screen "BWT Target Setpoints" 1280x800, template "Template"
   on GenerateScreen: "TitleUpdater"()
   Button "HmiScreenItemData_1" at 1,1 size 150x43; TextOn 'Back'; TextOff 'Commissioning'
      on Release: ActivateScreen("Commissioning Main Page", 0)
   AlarmView "Alarm view_1" at 0,777 size 1280x23
   IOField "I/O field_3" at 570,423 size 115x22; FormatPattern 9999.9; Unit Nm³/hr
      ProcessValue <- "2084_Setpoints_FIT420_LoLo"
   TextField "Text field_10" at 47,184 size 216x30; Text 'Description'
   TextField "Text field_6" at 579,184 size 100x30; Text 'Low Low'
   TextField "Text field_14" at 1099,184 size 100x30; Text 'High High'
   TextField "Text field_13" at 969,184 size 100x30; Text 'High'
   TextField "Text field_11" at 839,184 size 100x30; Text 'Setpoint'
   TextField "Text field_9" at 709,184 size 100x30; Text 'Low'
   IOField "I/O field_4" at 707,423 size 115x22; FormatPattern 9999.9; Unit Nm³/hr
      ProcessValue <- "2084_Setpoints_FIT420_Lo"
   IOField "I/O field_20" at 969,423 size 115x22; FormatPattern 9999.9; Unit Nm³/hr
      ProcessValue <- "2084_Setpoints_FIT420_Hi"
   IOField "I/O field_21" at 1099,423 size 115x22; FormatPattern 9999.9; Unit Nm³/hr
      ProcessValue <- "2084_Setpoints_FIT420_HiHi"
   TextField "Text field_8" at 295,184 size 100x30; Text 'Port'
   TextField "Text field_12" at 416,184 size 100x30; Text 'Starboard'
   IOField "I/O field_5" at 570,336 size 115x22; FormatPattern 9999.9; Unit Nm³/hr
      ProcessValue <- "2084_Setpoints_FIT418_LoLo"
   IOField "I/O field_29" at 707,336 size 115x22; FormatPattern 9999.9; Unit Nm³/hr
      ProcessValue <- "2084_Setpoints_FIT418_Lo"
   IOField "I/O field_39" at 969,336 size 115x22; FormatPattern 9999.9; Unit Nm³/hr
      ProcessValue <- "2084_Setpoints_FIT418_Hi"
   IOField "I/O field_40" at 1099,336 size 115x22; FormatPattern 9999.9; Unit Nm³/hr
      ProcessValue <- "2084_Setpoints_FIT418_HiHi"
   TextField "Text field_23" at 837,336 size 115x22; Text 'Text'
   TextField "Text field_24" at 837,423 size 115x22; Text 'Text'
   IOField "I/O field_19" at 837,624 size 115x22; FormatPattern 99.9; Unit  %
      ProcessValue <- "2084_Setpoints_DO_SP"
   TextField "Text field_34" at 47,624 size 220x22; Text 'DO428 DISOLVED OXYGEN'
   IOField "I/O field_36" at 295,624 size 115x22; FormatPattern 999.9; Unit %
      ProcessValue <- "20_TANKS_IP_DATA_RIO_02_FIRST_TANK_BWT_DO"
   IOField "I/O field_37" at 416,624 size 115x22; FormatPattern 999.9; Unit %
      ProcessValue <- "20_TANKS_IP_DATA_RIO_02_SECOND_TANK_BWT_DO"
   TextField "Text field_20" at 570,624 size 115x22; Text 'Text'
   TextField "Text field_30" at 707,624 size 115x22; Text 'Text'
   TextField "Text field_32" at 969,624 size 115x22; Text 'Text'
   TextField "Text field_36" at 1099,624 size 115x22; Text 'Text'
   TextField "Text field_35" at 47,579 size 220x22; Text 'PH426 PH LEVEL'
   IOField "I/O field_8" at 837,579 size 115x22; FormatPattern 9.9; Unit  ph
      ProcessValue <- "2084_Setpoints_PH_SP"
   IOField "I/O field_34" at 295,579 size 115x22; FormatPattern 9.9; Unit  ph
      ProcessValue <- "20_TANKS_IP_DATA_RIO_02_FIRST_TANK_BWT_PH"
   IOField "I/O field_35" at 416,579 size 115x22; FormatPattern 9.9; Unit  ph
      ProcessValue <- "20_TANKS_IP_DATA_RIO_02_SECOND_TANK_BWT_PH"
   TextField "Text field_19" at 570,579 size 115x22; Text 'Text'
   TextField "Text field_29" at 707,579 size 115x22; Text 'Text'
   TextField "Text field_31" at 969,579 size 115x22; Text 'Text'
   TextField "Text field_33" at 1099,579 size 115x22; Text 'Text'
   TextField "Text field_7" at 47,535 size 220x22; Text 'TT436 BWT TEMP'
   IOField "I/O field_38" at 1099,535 size 115x22; FormatPattern 999; Unit  DegC
      ProcessValue <- "2084_Setpoints_TT436_HiHi"
   IOField "I/O field_2" at 969,535 size 115x22; FormatPattern 999; Unit  DegC
      ProcessValue <- "2084_Setpoints_TT436_Hi"
   IOField "I/O field_32" at 295,535 size 115x22; FormatPattern 999.9; Unit  DegC
      ProcessValue <- "20_TANKS_IP_DATA_RIO_02_FIRST_TANK_BWT_TEMP"
   IOField "I/O field_33" at 416,535 size 115x22; FormatPattern 999.9; Unit  DegC
      ProcessValue <- "20_TANKS_IP_DATA_RIO_02_SECOND_TANK_BWT_TEMP"
   TextField "Text field_18" at 570,535 size 115x22; Text 'Text'
   TextField "Text field_26" at 837,535 size 115x22; Text 'Text'
   TextField "Text field_27" at 707,535 size 115x22; Text 'Text'
   TextField "Text field_5" at 47,490 size 220x22; Text 'LT422 BWT LEVEL'
   IOField "I/O field_6" at 969,490 size 115x22; Authorization "Parameter Change"; FormatPattern 999; Unit  %
      ProcessValue <- "2084_Setpoints_LT422_Hi"
   IOField "I/O field_11" at 707,490 size 115x22; Authorization "Parameter Change"; FormatPattern 999; Unit  %
      ProcessValue <- "2084_Setpoints_LT422_Lo"
   IOField "I/O field_30" at 295,490 size 115x22; FormatPattern s999.9; Unit %
      ProcessValue <- "20_TANKS_IP_DATA_RIO_02_FIRST_TANK_BWT_LEVEL"
   IOField "I/O field_31" at 416,490 size 115x22; FormatPattern s999.9; Unit %
      ProcessValue <- "20_TANKS_IP_DATA_RIO_02_SECOND_TANK_BWT_LEVEL"
   TextField "Text field_17" at 570,490 size 115x22; Text 'Text'
   TextField "Text field_25" at 837,490 size 115x22; Text 'Text'
   TextField "Text field_4" at 47,446 size 220x22; Text 'FIT 420 MBG FLOW'
   IOField "I/O field_28" at 358,446 size 115x22; FormatPattern 999.9; Unit Nm³/hr
      ProcessValue <- "20_TANKS_IP_DATA_RIO_02_FIRST_TANK_MBG_FLOW"
   TextField "Text field_16" at 47,401 size 220x22; Text 'FIT 419 MBG FLOW'
   IOField "I/O field_27" at 358,401 size 115x22; FormatPattern 999.9; Unit Nm³/hr
      ProcessValue <- "20_TANKS_IP_DATA_RIO_02_SECOND_TANK_MBG_FLOW"
   TextField "Text field_3" at 47,357 size 220x22; Text 'FIT418 USD FLOW'
   IOField "I/O field_25" at 358,357 size 115x22; FormatPattern 999.9; Unit Nm³/hr
      ProcessValue <- "20_TANKS_IP_DATA_RIO_02_FIRST_TANK_USD_FLOW"
   TextField "Text field_15" at 47,312 size 220x22; Text 'FIT417 USD FLOW'
   IOField "I/O field_23" at 358,312 size 115x22; FormatPattern 999.9; Unit Nm³/hr
      ProcessValue <- "20_TANKS_IP_DATA_RIO_02_SECOND_TANK_USD_FLOW"
   TextField "Text field_2" at 47,268 size 220x22; Text 'PT424 TANK PRESSURE'
   IOField "I/O field_15" at 570,268 size 115x22; FormatPattern 999.9; Unit  mBarg
      ProcessValue <- "2084_Setpoints_PIT424_LoLo"
   IOField "I/O field_17" at 1099,268 size 115x22; FormatPattern 999.9; Unit  mBarg
      ProcessValue <- "2084_Setpoints_PIT424_HiHi"
   IOField "I/O field_16" at 969,268 size 115x22; FormatPattern 999.9; Unit  mBarg
      ProcessValue <- "2084_Setpoints_PIT424_Hi"
   IOField "I/O field_14" at 707,268 size 115x22; FormatPattern 999.9; Unit  mBarg
      ProcessValue <- "2084_Setpoints_PIT424_Lo"
   IOField "I/O field_13" at 358,268 size 115x22; FormatPattern 999.9; Unit  mBarg
      ProcessValue <- "20_TANKS_IP_DATA_RIO_02_FIRST_TANK_TANKS_PRESS"
   TextField "Text field_22" at 837,268 size 115x22; Text 'Text'
   TextField "Text field_28" at 47,224 size 220x22; Text 'PT415 DECK IG PRESSURE'
   IOField "I/O field_9" at 570,224 size 115x22; FormatPattern 9.9; Unit  Barg
      ProcessValue <- "2084_Setpoints_PIT415_LoLo"
   IOField "I/O field_12" at 1099,224 size 115x22; FormatPattern 9.9; Unit  Barg
      ProcessValue <- "2084_Setpoints_PIT415_HiHi"
   IOField "I/O field_10" at 969,224 size 115x22; FormatPattern 9.9; Unit  Barg
      ProcessValue <- "2084_Setpoints_PIT415_Hi"
   IOField "I/O field_7" at 707,224 size 115x22; FormatPattern 9.9; Unit  Barg
      ProcessValue <- "2084_Setpoints_PIT415_Lo"
   IOField "I/O field_1" at 358,224 size 115x22; FormatPattern 9.9; Unit  Barg
      ProcessValue <- "20_TANKS_IP_DATA_RIO_02_FIRST_TANK_DECK_IG_PRESS"
   TextField "Text field_21" at 837,224 size 115x22; Text 'Text'
   TextField "Text field_1" at -7,151 size 450x30; Text 'BTCS TANK INSTRUMENT SETPOINTS'
   TextField "Text field_37" at 1099,490 size 115x22; Text 'Text'
   TextField "Text field_38" at 47,670 size 220x22; Text 'FIT 419 MBG FLOW PRESSURE SETPOINT'
   IOField "I/O field_18" at 358,670 size 115x22; FormatPattern 999.99; Unit BarG
      ProcessValue <- "21_FLOW_PRESSURE_SETPOINT_FIT_419_PRESSURE_SETPOINT"
   TextField "Text field_39" at 47,714 size 220x22; Text 'FIT 420 MBG FLOW PRESSURE SETPOINT'
   IOField "I/O field_22" at 358,714 size 115x22; FormatPattern 999.99; Unit BarG
      ProcessValue <- "21_FLOW_PRESSURE_SETPOINT_FIT_420_PRESSURE_SETPOINT"
   Group "Group" at 455,41 size 373x50
   Button "HmiScreenItemData_8" at 469,45 size 355x40; TextOn 'Back'; TextOff 'Text'
   TextField "Screen title" at 455,41 size 373x50; Text 'Screen title'

screen "BWT Process Times" 1280x800, template "Template"
   on GenerateScreen: "TitleUpdater"()
   Button "HmiScreenItemData_1" at 1,1 size 150x43; TextOn 'Back'; TextOff 'Commissioning'
      on Release: ActivateScreen("Commissioning Main Page", 0)
   Button "Button_1" at 21,736 size 161x32; TextOff 'IGG Step Times'
      on Activate: ActivateScreen("IGG Max Step Times", 0)
   Button "Button_2" at 1091,736 size 161x32; TextOff 'BC Step Times'
      on Activate: ActivateScreen("BC Max Step Times", 0)
   AlarmView "Alarm view_1" at 0,777 size 1280x23
   TextField "Text field_29" at 345,95 size 65x20; Text 'Time (s)'
   TextField "Text field_65" at 40,120 size 300x25; Text 'DE-OX PRE-GTT OPEN DELAY'
   TextField "Text field_42" at 40,95 size 89x20; Text 'Description'
   IOField "I/O field_128" at 345,120 size 65x25; Authorization "Parameter Change"; FormatPattern 999
      ProcessValue <- "2086_Times_DEOX_PRE_GTT_OPN_DLY"
   TextField "Text field_53" at 40,66 size 197x26; Text 'BWT Process Times'
   TextField "Text field_1" at 40,150 size 300x25; Text 'DE-OX POST-GTT CLOSE DELAY'
   IOField "I/O field_1" at 345,150 size 65x25; Authorization "Parameter Change"; FormatPattern 999
      ProcessValue <- "2086_Times_DEOX_PRE_GTT_CLS_DLY"
   TextField "Text field_2" at 40,180 size 300x25; Text 'RE-OX PRE-GTT OPEN DELAY'
   IOField "I/O field_2" at 345,180 size 65x25; Authorization "Parameter Change"; FormatPattern 999
      ProcessValue <- "2086_Times_REOX_PRE_GTT_OPN_DLY"
   TextField "Text field_3" at 40,210 size 300x25; Text 'RE-OX POST-GTT CLOSE DELAY'
   IOField "I/O field_3" at 345,210 size 65x25; Authorization "Parameter Change"; FormatPattern 999
      ProcessValue <- "2086_Times_REOX_PRE_GTT_CLS_DLY"
   TextField "Text field_8" at 775,95 size 65x20; Text 'Time (s)'
   TextField "Text field_9" at 40,240 size 300x25; Text 'AT DE-OX CONFIRMATION TIME'
   TextField "Text field_10" at 470,95 size 89x20; Text 'Description'
   IOField "I/O field_8" at 345,240 size 65x25; Authorization "Parameter Change"; FormatPattern 999
      ProcessValue <- "2086_Times_AT_DEOX_CNF_TIME"
   TextField "Text field_11" at 40,270 size 300x25; Text 'AT RE-OX CONFIRMATION TIME'
   IOField "I/O field_9" at 345,270 size 65x25; Authorization "Parameter Change"; FormatPattern 999
      ProcessValue <- "2086_Times_AT_REOX_CNF_TIME"
   TextField "Text field_4" at 894,120 size 300x25; Text 'VOYAGE TIME REMAINING POPUP REAPPEAR'
   IOField "I/O field_4" at 1199,120 size 65x25; Authorization "Parameter Change"; FormatPattern 999; Unit h
      ProcessValue <- "2086_Times_Stage Warning"
   TextField "Text field_5" at 1176,95 size 88x20; Text 'Time (secs)'
   TextField "Text field_6" at 894,95 size 89x20; Text 'Description'
   TextField "Text field_13" at 471,120 size 300x25; Text 'TT426PORT Alarm Delay'
   IOField "I/O field_7" at 776,120 size 65x25; Authorization "Parameter Change"; FormatPattern 999
      ProcessValue <- "2086_Times_TT426_PORT_Alarm Delay"
   TextField "Text field_14" at 471,150 size 300x25; Text 'TT426STAR Alarm Delay'
   IOField "I/O field_10" at 776,150 size 65x25; Authorization "Parameter Change"; FormatPattern 999
      ProcessValue <- "2086_Times_TT426_STAR_Alarm Delay"
   TextField "Text field_15" at 471,180 size 300x25; Text 'FIT418PORT Alarm Delay'
   IOField "I/O field_11" at 776,180 size 65x25; Authorization "Parameter Change"; FormatPattern 999
      ProcessValue <- "2086_Times_FIT418PORT Alarm Delay"
   TextField "Text field_16" at 471,210 size 300x25; Text 'FIT420PORT Alarm Delay'
   IOField "I/O field_12" at 776,210 size 65x25; Authorization "Parameter Change"; FormatPattern 999
      ProcessValue <- "2086_Times_FIT420PORT Alarm Delay"
   TextField "Text field_17" at 471,240 size 300x25; Text 'FIT417STAR Alarm Delay'
   IOField "I/O field_13" at 776,240 size 65x25; Authorization "Parameter Change"; FormatPattern 999
      ProcessValue <- "2086_Times_FIT417STAR Alarm Delay"
   TextField "Text field_18" at 470,270 size 300x25; Text 'FIT419STAR Alarm Delay'
   IOField "I/O field_14" at 775,270 size 65x25; Authorization "Parameter Change"; FormatPattern 999
      ProcessValue <- "2086_Times_FIT419STAR Alarm Delay"
   TextField "Text field_19" at 470,300 size 300x25; Text 'PT415PORT Alarm Delay'
   IOField "I/O field_15" at 775,300 size 65x25; Authorization "Parameter Change"; FormatPattern 999
      ProcessValue <- "2086_Times_PT415 Alarm Delay"
   TextField "Text field_20" at 470,331 size 300x25; Text 'PT424PORT Alarm Delay'
   IOField "I/O field_16" at 775,331 size 65x25; Authorization "Parameter Change"; FormatPattern 999
      ProcessValue <- "2086_Times_PIT424 Alarm Delay"
   TextField "Text field_21" at 470,362 size 300x25; Text 'LS425PORT Alarm Delay'
   IOField "I/O field_17" at 775,362 size 65x25; Authorization "Parameter Change"; FormatPattern 999
      ProcessValue <- "2086_Times_LS425 Port Alarm Delay"
   TextField "Text field_22" at 470,393 size 300x25; Text 'LS425STAR Alarm Delay'
   IOField "I/O field_18" at 775,393 size 65x25; Authorization "Parameter Change"; FormatPattern 999
      ProcessValue <- "2086_Times_LS425 Star Alarm Delay"
   TextField "Text field_23" at 470,424 size 300x25; Text 'PS436 Alarm Delay'
   IOField "I/O field_19" at 775,424 size 65x25; Authorization "Parameter Change"; FormatPattern 999
      ProcessValue <- "2086_Times_PS436 Alarm Delay"
   Group "Group" at 455,41 size 373x50
   TextField "Text field_7" at 470,456 size 300x25; Text 'Tank Alarm Reset Time'
   IOField "I/O field_5" at 775,456 size 65x25; Authorization "Parameter Change"; FormatPattern 999
      ProcessValue <- "2086_Times_Tank Alarm Reset Time"
   TextField "Text field_12" at 470,488 size 300x25; Text 'Alarm Enable Delay'
   IOField "I/O field_6" at 775,488 size 65x25; Authorization "Parameter Change"; FormatPattern 999
      ProcessValue <- "2086_Times_Alarm Enable Delay"
   TextField "Text field_24" at 894,150 size 300x25; Text 'CV422 FPT Maximum Travel Time'
   IOField "I/O field_20" at 1199,150 size 65x25; Authorization "Parameter Change"; FormatPattern 999
      ProcessValue <- "2086_Times_CV422_FPT_MAX_TRVL_TIME"
   TextField "Text field_25" at 894,181 size 300x25; Text 'CV422 1P Maximum Travel Time'
   IOField "I/O field_21" at 1199,181 size 65x25; Authorization "Parameter Change"; FormatPattern 999
      ProcessValue <- "2086_Times_CV422_1P_MAX_TRVL_TIME"
   TextField "Text field_26" at 894,211 size 300x25; Text 'CV421 1S Maximum Travel Time'
   IOField "I/O field_22" at 1199,211 size 65x25; Authorization "Parameter Change"; FormatPattern 999
      ProcessValue <- "2086_Times_CV421_1S_MAX_TRVL_TIME"
   TextField "Text field_27" at 894,242 size 300x25; Text 'CV422 2P Maximum Travel Time'
   IOField "I/O field_23" at 1199,242 size 65x25; Authorization "Parameter Change"; FormatPattern 999
      ProcessValue <- "2086_Times_CV422_2P_MAX_TRVL_TIME"
   TextField "Text field_28" at 894,273 size 300x25; Text 'CV421 2S Maximum Travel Time'
   IOField "I/O field_24" at 1199,273 size 65x25; Authorization "Parameter Change"; FormatPattern 999
      ProcessValue <- "2086_Times_CV421_2S_MAX_TRVL_TIME"
   TextField "Text field_30" at 894,303 size 300x25; Text 'CV422 3P Maximum Travel Time'
   IOField "I/O field_25" at 1199,303 size 65x25; Authorization "Parameter Change"; FormatPattern 999
      ProcessValue <- "2086_Times_CV422_3P_MAX_TRVL_TIME"
   TextField "Text field_31" at 894,334 size 300x25; Text 'CV421 3S Maximum Travel Time'
   IOField "I/O field_26" at 1199,334 size 65x25; Authorization "Parameter Change"; FormatPattern 999
      ProcessValue <- "2086_Times_CV421_3S_MAX_TRVL_TIME"
   TextField "Text field_32" at 894,365 size 300x25; Text 'CV422 4P Maximum Travel Time'
   IOField "I/O field_27" at 1199,365 size 65x25; Authorization "Parameter Change"; FormatPattern 999
      ProcessValue <- "2086_Times_CV422_4P_MAX_TRVL_TIME"
   TextField "Text field_33" at 894,396 size 300x25; Text 'CV421 4S Maximum Travel Time'
   IOField "I/O field_28" at 1199,396 size 65x25; Authorization "Parameter Change"; FormatPattern 999
      ProcessValue <- "2086_Times_CV421_4S_MAX_TRVL_TIME"
   TextField "Text field_34" at 894,426 size 300x25; Text 'CV422 5P Maximum Travel Time'
   IOField "I/O field_29" at 1199,426 size 65x25; Authorization "Parameter Change"; FormatPattern 999
      ProcessValue <- "2086_Times_CV422_5P_MAX_TRVL_TIME"
   TextField "Text field_35" at 894,457 size 300x25; Text 'CV421 5S Maximum Travel Time'
   IOField "I/O field_30" at 1199,457 size 65x25; Authorization "Parameter Change"; FormatPattern 999
      ProcessValue <- "2086_Times_CV421_5S_MAX_TRVL_TIME"
   TextField "Text field_36" at 894,488 size 300x25; Text 'CV422 6P Maximum Travel Time'
   IOField "I/O field_31" at 1199,488 size 65x25; Authorization "Parameter Change"; FormatPattern 999
      ProcessValue <- "2086_Times_CV422_6P_MAX_TRVL_TIME"
   TextField "Text field_37" at 894,519 size 300x25; Text 'CV421 6S Maximum Travel Time'
   IOField "I/O field_32" at 1198,519 size 65x25; Authorization "Parameter Change"; FormatPattern 999
      ProcessValue <- "2086_Times_CV421_6S_MAX_TRVL_TIME"
   TextField "Text field_38" at 893,550 size 300x25; Text 'CV421 APT Maximum Travel Time'
   IOField "I/O field_33" at 1197,550 size 65x25; Authorization "Parameter Change"; FormatPattern 999
      ProcessValue <- "2086_Times_CV422_APT_MAX_TRVL_TIME"
   Button "HmiScreenItemData_8" at 469,45 size 355x40; TextOn 'Back'; TextOff 'Text'
   TextField "Screen title" at 455,41 size 373x50; Text 'Screen title'

screen "GCU Digital Outputs" 1280x800, template "Template"
   on GenerateScreen: "TitleUpdater"()
   Button "HmiScreenItemData_1" at 1,1 size 150x43; TextOn 'Back'; TextOff 'Commissioning'
      on Release: ActivateScreen("Commissioning Main Page", 0)
   AlarmView "Alarm view_1" at 0,777 size 1280x23
   Button "Button_19" at 187,97 size 70x30; TextOff 'Override'
      on Press: InvertBit("80_From_HMI_MAN_DQ_136_0")
      Visibility <- "82_To_HMI_CRNT_MODE_GCU"
      Appearance <- "80_From_HMI_MAN_DQ_136_0"
   TextField "Text field_2" at 165,42 size 300x30; Text 'GCU Control PLC (Rack 3)'
   TextField "Text field_34" at 725,72 size 60x30; Text 'Q 2'
   TextField "Text field_35" at 725,382 size 70x22; Text 'Q 138.7'
   Circle "Circle_16" at 811,382 size 20x20
      Appearance <- "14_DQ_DATA_R3_SPR_DQ_138_7"
   TextField "Text field_36" at 845,382 size 230x22; Text 'R3_SPR_DQ_138_7'
   TextField "Text field_39" at 725,342 size 70x22; Text 'Q 138.6'
   Circle "Circle_17" at 811,342 size 20x20
      Appearance <- "14_DQ_DATA_CV_421_3S"
   TextField "Text field_40" at 845,342 size 230x22; Text 'CV421 GTT 3 STBD'
   TextField "Text field_41" at 725,302 size 70x22; Text 'Q 138.5'
   Circle "Circle_18" at 811,302 size 20x20
      Appearance <- "14_DQ_DATA_CV_422_3P"
   TextField "Text field_42" at 845,302 size 230x22; Text 'CV422 GTT 3 PORT'
   TextField "Text field_43" at 725,262 size 70x22; Text 'Q 138.4'
   Circle "Circle_19" at 811,262 size 20x20
      Appearance <- "14_DQ_DATA_CV_421_2S"
   TextField "Text field_44" at 845,262 size 230x22; Text 'CV421 GTT 2 STBD'
   TextField "Text field_45" at 725,222 size 70x22; Text 'Q 138.3'
   Circle "Circle_20" at 811,222 size 20x20
      Appearance <- "14_DQ_DATA_CV_422_2P"
   TextField "Text field_46" at 845,222 size 230x22; Text 'CV422 GTT 2 PORT'
   TextField "Text field_47" at 725,182 size 70x22; Text 'Q 138.2'
   Circle "Circle_21" at 811,182 size 20x20
      Appearance <- "14_DQ_DATA_CV_421_1S"
   TextField "Text field_48" at 845,182 size 230x22; Text 'CV421 GTT 1 STBD'
   TextField "Text field_49" at 725,142 size 70x22; Text 'Q 138.1'
   Circle "Circle_22" at 811,142 size 20x20
      Appearance <- "14_DQ_DATA_CV_422_1P"
   TextField "Text field_50" at 845,142 size 230x22; Text 'CV422 GTT 1 PORT'
   TextField "Text field_51" at 725,102 size 70x22; Text 'Q 138.0'
   Circle "Circle_23" at 811,102 size 20x20
      Appearance <- "14_DQ_DATA_CV_422_FPT"
   TextField "Text field_52" at 845,102 size 230x22; Text 'CV422 GTT FPT'
   TextField "Text field_3" at 269,72 size 60x30; Text 'Q 0'
   TextField "Text field_15" at 269,382 size 70x22; Text 'Q 136.7'
   Circle "Circle_7" at 354,382 size 20x20
      Appearance <- "10_DI_DATA_E_400_RUN"
   TextField "Text field_16" at 389,382 size 230x22; Text 'E400 PGC START'
   TextField "Text field_13" at 269,342 size 70x22; Text 'Q 136.6'
   Circle "Circle_6" at 354,342 size 20x20
      Appearance <- "10_DI_DATA_CV406_OPN"
   TextField "Text field_14" at 389,342 size 230x22; Text 'CV406 GAS TO DECK'
   TextField "Text field_11" at 269,302 size 70x22; Text 'Q 136.5'
   Circle "Circle_5" at 354,302 size 20x20
      Appearance <- "10_DI_DATA_CV441_CLSD"
   TextField "Text field_12" at 389,302 size 230x22; Text 'CV441 AMBIENT AIR'
   TextField "Text field_4" at 269,262 size 70x22; Text 'Q 136.4'
   Circle "Circle_4" at 354,262 size 20x20
      Appearance <- "10_DI_DATA_CV411_OPN"
   TextField "Text field_10" at 389,262 size 230x22; Text 'CV411 BLOCK VALVE 2'
   TextField "Text field_7" at 269,222 size 70x22; Text 'Q 136.3'
   Circle "Circle_3" at 354,222 size 20x20
      Appearance <- "10_DI_DATA_CV409_CLSD"
   TextField "Text field_8" at 389,222 size 230x22; Text 'CV409 BLEED VALVE'
   TextField "Text field_5" at 269,182 size 70x22; Text 'Q 136.2'
   Circle "Circle_2" at 354,182 size 20x20
      Appearance <- "10_DI_DATA_CV407_OPN"
   TextField "Text field_6" at 389,182 size 230x22; Text 'CV407 BLOCK VALVE 1'
   TextField "Text field_17" at 269,142 size 70x22; Text 'Q 136.1'
   Circle "Circle_1" at 354,142 size 20x20
      Appearance <- "10_DI_DATA_CV341_CLSD"
   TextField "Text field_18" at 389,142 size 230x22; Text 'CV341 DRAIN VALVE'
   TextField "Text field_38" at 269,102 size 70x22; Text 'Q 136.0'
   Circle "Circle_33" at 354,102 size 20x20
      Appearance <- "10_DI_DATA_CV358_OPN"
   TextField "Text field_19" at 389,102 size 230x22; Text 'CV358 FCW FILL VALVE'
   TextField "Text field_53" at 725,422 size 60x30; Text 'Q 3'
   TextField "Text field_54" at 725,732 size 70x22; Text 'Q 139.7'
   Circle "Circle_24" at 811,732 size 20x20
      Appearance <- "14_DQ_DATA_R3_SPR_DQ_139_7"
   TextField "Text field_55" at 845,732 size 230x22; Text 'R3_SPR_DQ_139_7'
   TextField "Text field_56" at 725,692 size 70x22; Text 'Q 139.6'
   Circle "Circle_25" at 811,692 size 20x20
      Appearance <- "14_DQ_DATA_CV_422_APT"
   TextField "Text field_57" at 845,692 size 230x22; Text 'CV422 GTT APT'
   TextField "Text field_58" at 725,652 size 70x22; Text 'Q 139.5'
   Circle "Circle_26" at 811,652 size 20x20
      Appearance <- "14_DQ_DATA_CV_421_6S"
   TextField "Text field_60" at 725,612 size 70x22; Text 'Q 139.4'
   Circle "Circle_27" at 811,612 size 20x20
      Appearance <- "14_DQ_DATA_CV_422_6P"
   TextField "Text field_62" at 725,572 size 70x22; Text 'Q 139.3'
   Circle "Circle_28" at 811,572 size 20x20
      Appearance <- "14_DQ_DATA_CV_421_5S"
   TextField "Text field_64" at 725,532 size 70x22; Text 'Q 139.2'
   Circle "Circle_29" at 811,532 size 20x20
      Appearance <- "14_DQ_DATA_CV_422_5P"
   TextField "Text field_66" at 725,492 size 70x22; Text 'Q 139.1'
   Circle "Circle_30" at 811,492 size 20x20
      Appearance <- "14_DQ_DATA_CV_421_4S"
   TextField "Text field_68" at 725,452 size 70x22; Text 'Q 139.0'
   Circle "Circle_31" at 811,452 size 20x20
      Appearance <- "14_DQ_DATA_CV_422_4P"
   TextField "Text field_20" at 269,422 size 60x30; Text 'Q 1'
   TextField "Text field_21" at 269,732 size 70x22; Text 'Q 137.7'
   Circle "Circle_8" at 354,732 size 20x20
      Appearance <- "14_DQ_DATA_E_400_STP"
   TextField "Text field_22" at 389,732 size 230x22; Text 'E400 PGC STOP'
   TextField "Text field_23" at 269,692 size 70x22; Text 'Q 137.6'
   Circle "Circle_9" at 354,692 size 20x20
      Appearance <- "14_DQ_DATA_13P5"
   TextField "Text field_24" at 389,692 size 230x22; Text '13P5 BUZZER'
   TextField "Text field_25" at 269,652 size 70x22; Text 'Q 137.5'
   Circle "Circle_10" at 354,652 size 20x20
      Appearance <- "14_DQ_DATA_13P4"
   TextField "Text field_26" at 389,652 size 230x22; Text '13P4 BALLAST HiHi'
   TextField "Text field_27" at 269,612 size 70x22; Text 'Q 137.4'
   Circle "Circle_11" at 354,612 size 20x20
      Appearance <- "14_DQ_DATA_13P3"
   TextField "Text field_28" at 389,612 size 230x22; Text '13P3 RUNNING'
   TextField "Text field_29" at 269,572 size 70x22; Text 'Q 137.3'
   Circle "Circle_12" at 354,572 size 20x20
      Appearance <- "14_DQ_DATA_13P2"
   TextField "Text field_30" at 389,572 size 230x22; Text '13P2 ALARM'
   TextField "Text field_31" at 269,532 size 70x22; Text 'Q 137.2'
   Circle "Circle_13" at 354,532 size 20x20
      Appearance <- "14_DQ_DATA_13P1"
   TextField "Text field_32" at 389,532 size 230x22; Text '13P1 WARNING'
   TextField "Text field_33" at 269,492 size 70x22; Text 'Q 137.1'
   Circle "Circle_14" at 354,492 size 20x20
      Appearance <- "14_DQ_DATA_P_304"
   TextField "Text field_37" at 389,492 size 230x22; Text 'P304 BOOSTER PUMP'
   TextField "Text field_70" at 269,452 size 70x22; Text 'Q 137.0'
   Circle "Circle_15" at 354,452 size 20x20
      Appearance <- "14_DQ_DATA_P_303"
   TextField "Text field_71" at 389,452 size 230x22; Text 'P303 RECIRC PUMP'
   TextField "Text field_59" at 845,652 size 230x22; Text 'CV421 GTT 6 STBD'
   TextField "Text field_61" at 845,612 size 230x22; Text 'CV422 GTT 6 PORT'
   TextField "Text field_63" at 845,572 size 230x22; Text 'CV421 GTT 5 STBD'
   TextField "Text field_65" at 845,532 size 230x22; Text 'CV422 GTT 5 PORT'
   TextField "Text field_67" at 845,492 size 230x22; Text 'CV421 GTT 4 STBD'
   TextField "Text field_69" at 845,452 size 230x22; Text 'CV422 GTT 4 PORT'
   Button "Button_1" at 647,98 size 70x30; TextOff 'Override'
      on Press: InvertBit("80_From_HMI_MAN_DQ_138_0")
      Visibility <- "82_To_HMI_CRNT_MODE_GCU"
      Appearance <- "80_From_HMI_MAN_DQ_138_0"
   Button "Button_2" at 187,137 size 70x30; TextOff 'Override'
      on Press: InvertBit("80_From_HMI_MAN_DQ_136_1")
      Visibility <- "82_To_HMI_CRNT_MODE_GCU"
      Appearance <- "80_From_HMI_MAN_DQ_136_1"
   Button "Button_3" at 187,177 size 70x30; TextOff 'Override'
      on Press: InvertBit("80_From_HMI_MAN_DQ_136_2")
      Visibility <- "82_To_HMI_CRNT_MODE_GCU"
      Appearance <- "80_From_HMI_MAN_DQ_136_2"
   Button "Button_4" at 187,217 size 70x30; TextOff 'Override'
      on Press: InvertBit("80_From_HMI_MAN_DQ_136_3")
      Visibility <- "82_To_HMI_CRNT_MODE_GCU"
      Appearance <- "80_From_HMI_MAN_DQ_136_3"
   Button "Button_5" at 187,257 size 70x30; TextOff 'Override'
      on Press: InvertBit("80_From_HMI_MAN_DQ_136_4")
      Visibility <- "82_To_HMI_CRNT_MODE_GCU"
      Appearance <- "80_From_HMI_MAN_DQ_136_4"
   Button "Button_6" at 187,297 size 70x30; TextOff 'Override'
      on Press: InvertBit("80_From_HMI_MAN_DQ_136_5")
      Visibility <- "82_To_HMI_CRNT_MODE_GCU"
      Appearance <- "80_From_HMI_MAN_DQ_136_5"
   Button "Button_7" at 187,337 size 70x30; TextOff 'Override'
      on Press: InvertBit("80_From_HMI_MAN_DQ_136_6")
      Visibility <- "82_To_HMI_CRNT_MODE_GCU"
      Appearance <- "80_From_HMI_MAN_DQ_136_6"
   Button "Button_8" at 187,377 size 70x30; TextOff 'Override'
      on Press: InvertBit("80_From_HMI_MAN_DQ_136_7")
      Visibility <- "82_To_HMI_CRNT_MODE_GCU"
      Appearance <- "80_From_HMI_MAN_DQ_136_7"
   Button "Button_10" at 187,447 size 70x30; TextOff 'Override'
      on Press: InvertBit("80_From_HMI_MAN_DQ_137_0")
      Visibility <- "82_To_HMI_CRNT_MODE_GCU"
      Appearance <- "80_From_HMI_MAN_DQ_137_0"
   Button "Button_9" at 187,487 size 70x30; TextOff 'Override'
      on Press: InvertBit("80_From_HMI_MAN_DQ_137_1")
      Visibility <- "82_To_HMI_CRNT_MODE_GCU"
      Appearance <- "80_From_HMI_MAN_DQ_137_1"
   Button "Button_11" at 187,527 size 70x30; TextOff 'Override'
      on Press: InvertBit("80_From_HMI_MAN_DQ_137_2")
      Visibility <- "82_To_HMI_CRNT_MODE_GCU"
      Appearance <- "80_From_HMI_MAN_DQ_137_2"
   Button "Button_12" at 187,567 size 70x30; TextOff 'Override'
      on Press: InvertBit("80_From_HMI_MAN_DQ_137_3")
      Visibility <- "82_To_HMI_CRNT_MODE_GCU"
      Appearance <- "80_From_HMI_MAN_DQ_137_3"
   Button "Button_13" at 187,607 size 70x30; TextOff 'Override'
      on Press: InvertBit("80_From_HMI_MAN_DQ_137_4")
      Visibility <- "82_To_HMI_CRNT_MODE_GCU"
      Appearance <- "80_From_HMI_MAN_DQ_137_4"
   Button "Button_14" at 187,647 size 70x30; TextOff 'Override'
      on Press: InvertBit("80_From_HMI_MAN_DQ_137_5")
      Visibility <- "82_To_HMI_CRNT_MODE_GCU"
      Appearance <- "80_From_HMI_MAN_DQ_137_5"
   Button "Button_15" at 187,687 size 70x30; TextOff 'Override'
      on Press: InvertBit("80_From_HMI_MAN_DQ_137_6")
      Visibility <- "82_To_HMI_CRNT_MODE_GCU"
      Appearance <- "80_From_HMI_MAN_DQ_137_6"
   Button "Button_16" at 187,727 size 70x30; TextOff 'Override'
      on Press: InvertBit("80_From_HMI_MAN_DQ_137_7")
      Visibility <- "82_To_HMI_CRNT_MODE_GCU"
      Appearance <- "80_From_HMI_MAN_DQ_137_7"
   Button "Button_17" at 647,138 size 70x30; TextOff 'Override'
      on Press: InvertBit("80_From_HMI_MAN_DQ_138_1")
      Visibility <- "82_To_HMI_CRNT_MODE_GCU"
      Appearance <- "80_From_HMI_MAN_DQ_138_1"
   Button "Button_18" at 647,178 size 70x30; TextOff 'Override'
      on Press: InvertBit("80_From_HMI_MAN_DQ_138_2")
      Visibility <- "82_To_HMI_CRNT_MODE_GCU"
      Appearance <- "80_From_HMI_MAN_DQ_138_2"
   Button "Button_20" at 647,218 size 70x30; TextOff 'Override'
      on Press: InvertBit("80_From_HMI_MAN_DQ_138_3")
      Visibility <- "82_To_HMI_CRNT_MODE_GCU"
      Appearance <- "80_From_HMI_MAN_DQ_138_3"
   Button "Button_21" at 647,258 size 70x30; TextOff 'Override'
      on Press: InvertBit("80_From_HMI_MAN_DQ_138_4")
      Visibility <- "82_To_HMI_CRNT_MODE_GCU"
      Appearance <- "80_From_HMI_MAN_DQ_138_4"
   Button "Button_22" at 647,298 size 70x30; TextOff 'Override'
      on Press: InvertBit("80_From_HMI_MAN_DQ_138_5")
      Visibility <- "82_To_HMI_CRNT_MODE_GCU"
      Appearance <- "80_From_HMI_MAN_DQ_138_5"
   Button "Button_23" at 647,338 size 70x30; TextOff 'Override'
      on Press: InvertBit("80_From_HMI_MAN_DQ_138_6")
      Visibility <- "82_To_HMI_CRNT_MODE_GCU"
      Appearance <- "80_From_HMI_MAN_DQ_138_6"
   Button "Button_24" at 647,378 size 70x30; TextOff 'Override'
      on Press: InvertBit("80_From_HMI_MAN_DQ_138_7")
      Visibility <- "82_To_HMI_CRNT_MODE_GCU"
      Appearance <- "80_From_HMI_MAN_DQ_138_7"
   Button "Button_25" at 647,448 size 70x30; TextOff 'Override'
      on Press: InvertBit("80_From_HMI_MAN_DQ_139_0")
      Visibility <- "82_To_HMI_CRNT_MODE_GCU"
      Appearance <- "80_From_HMI_MAN_DQ_139_0"
   Button "Button_26" at 647,488 size 70x30; TextOff 'Override'
      on Press: InvertBit("80_From_HMI_MAN_DQ_139_1")
      Visibility <- "82_To_HMI_CRNT_MODE_GCU"
      Appearance <- "80_From_HMI_MAN_DQ_139_1"
   Button "Button_27" at 647,528 size 70x30; TextOff 'Override'
      on Press: InvertBit("80_From_HMI_MAN_DQ_139_2")
      Visibility <- "82_To_HMI_CRNT_MODE_GCU"
      Appearance <- "80_From_HMI_MAN_DQ_139_2"
   Button "Button_28" at 647,568 size 70x30; TextOff 'Override'
      on Press: InvertBit("80_From_HMI_MAN_DQ_139_3")
      Visibility <- "82_To_HMI_CRNT_MODE_GCU"
      Appearance <- "80_From_HMI_MAN_DQ_139_3"
   Button "Button_29" at 647,608 size 70x30; TextOff 'Override'
      on Press: InvertBit("80_From_HMI_MAN_DQ_139_4")
      Visibility <- "82_To_HMI_CRNT_MODE_GCU"
      Appearance <- "80_From_HMI_MAN_DQ_139_4"
   Button "Button_30" at 647,648 size 70x30; TextOff 'Override'
      on Press: InvertBit("80_From_HMI_MAN_DQ_139_5")
      Visibility <- "82_To_HMI_CRNT_MODE_GCU"
      Appearance <- "80_From_HMI_MAN_DQ_139_5"
   Button "Button_31" at 647,688 size 70x30; TextOff 'Override'
      on Press: InvertBit("80_From_HMI_MAN_DQ_139_6")
      Visibility <- "82_To_HMI_CRNT_MODE_GCU"
      Appearance <- "80_From_HMI_MAN_DQ_139_6"
   Button "Button_32" at 647,728 size 70x30; TextOff 'Override'
      on Press: InvertBit("80_From_HMI_MAN_DQ_139_7")
      Visibility <- "82_To_HMI_CRNT_MODE_GCU"
      Appearance <- "80_From_HMI_MAN_DQ_139_7"
   Group "Group" at 852,44 size 373x50
   Button "HmiScreenItemData_8" at 866,48 size 355x40; TextOn 'Back'; TextOff 'Text'
   TextField "Screen title" at 852,44 size 373x50; Text 'Screen title'

PopupScreen "Voyage Time Warning" 665x250
   Button "Button_1" at 0,0 size 665x250; TextOff 'Voyage Time Insufficient, Minimum Voyage Time For Treatment Is Days.'
      on Release: ActivateScreen("Balast Water Treatment Setup", 0)
   IOField "I/O field_1" at 359,124 size 82x50; FormatPattern 999
      ProcessValue <- "2102_TIME_CALCS_DB_TOT_SEQ_DAYS"
   Button "Button_2" at 208,187 size 250x35; TextOff 'OK, Adjust Voyage Time'
      on Release: ActivateScreen("Balast Water Treatment Setup", 0); function_efd93a16("Voyage Time Warning", 0, 0, -1, -1, 1)

PopupScreen "Treatment Cycle Completed" 665x230
   Button "Button_1" at 0,0 size 665x230; TextOff 'TREATMENT CYCLE COMPLETED'
      on Click: function_efd93a16("Treatment Cycle Completed", 0, 0, -1, -1, 1)

screen "Balast Water Treatment Setup" 1280x800, template "Template"
   Button "HmiScreenItemData_1" at 1,1 size 150x40; TextOn 'Back'; TextOff 'Main Index'
      on Release: ActivateScreen("02 Main Index", 0)
   Button "HmiScreenItemData_8" at 276,83 size 219x27; TextOn 'Back'; TextOff 'Plant Operation'
   Button "HmiScreenItemData_23" at 282,116 size 150x47; TextOn 'Back'; TextOff 'Accept & Launch'; Authorization "Operating Mode"
      Appearance <- "2110_BTCS_CNTRL_DB_BTCS_STATE"
      on Release: function_efd93a16("BWTS Start Confirm", 400, 200, -1, -1, 1)
      ObjectEnable <- "82_To_HMI_CRNT_MODE_GCU"
   Button "HmiScreenItemData_14" at 828,54 size 416x27; TextOn 'Back'; TextOff 'Treatment Durations'
   TextField "Text field_1" at 925,535 size 220x18; Text 'Tank Water Low Level (LT421)'
   TextField "Text field_2" at 925,573 size 220x18; Text 'Tank Water Low Level (LT422)'
   TextField "Text field_3" at 925,501 size 85x18; Text 'Description'
   TextField "Text field_5" at 925,611 size 215x18; Text 'De-Oxygenation DO Set Point'
   TextField "Text field_6" at 1164,501 size 67x18; Text 'Setpoint'
   Button "HmiScreenItemData_15" at 915,461 size 329x27; TextOn 'Back'; TextOff 'Ballast Tank Treatment Settings'
   IOField "I/O field_4" at 1153,530 size 80x28; Authorization "Operate"; FormatPattern 999.9; Unit  %
      ProcessValue <- "2084_Setpoints_LT421_Lo"
   IOField "I/O field_5" at 1153,568 size 80x28; Authorization "Operate"; FormatPattern 999.9; Unit  %
      ProcessValue <- "2084_Setpoints_LT422_Lo"
   IOField "I/O field_6" at 1153,606 size 80x28; Authorization "Operate"; FormatPattern 99.9; Unit  mg/l
      ProcessValue <- "2084_Setpoints_DO_SP"
   Button "HmiScreenItemData_16" at 482,461 size 334x27; TextOn 'Back'; TextOff 'Manual Ballast Tank Selection'
   Button "HmiScreenItemData_34" at 43,83 size 230x27; TextOn 'Back'; TextOff 'Plant Mode of Operation'
   Button "HmiScreenItemData_18" at 43,54 size 452x27; TextOn 'Back'; TextOff 'Ballast Water Treatment'
   Button "HmiScreenItemData_40" at 508,54 size 300x27; TextOn 'Back'; TextOff 'Treatment Status'
   TextField "Text field_14" at 837,94 size 85x18; Text 'Description'
   TextField "Text field_17" at 1054,94 size 67x18; Text 'Setpoint'
   IOField "I/O field_10" at 1040,132 size 92x27; Authorization "Operating Mode"; FormatPattern 999.99; Unit  Days
      ProcessValue <- "2115_VOYAGE_TIME_DAYS_VOYAGE_DAYS"
   IOField "I/O field_12" at 1040,267 size 79x28; Authorization "Commissioning"; FormatPattern 999; Unit  Hrs
      ProcessValue <- "2110_BTCS_CNTRL_DB_DE_OX_HRS"
   IOField "I/O field_13" at 1040,335 size 79x28; Authorization "Commissioning"; FormatPattern 999; Unit  Hrs
      ProcessValue <- "2110_BTCS_CNTRL_DB_DWELL_HRS"
   IOField "I/O field_14" at 1040,369 size 79x28; Authorization "Commissioning"; FormatPattern 999; Unit  Hrs
      ProcessValue <- "2110_BTCS_CNTRL_DB_RE_OX_HRS"
   IOField "I/O field_15" at 1040,403 size 79x28; Authorization "Commissioning"; FormatPattern 999; Unit  Hrs
      ProcessValue <- "2110_BTCS_CNTRL_DB_POST_DWELL_HRS"
   Button "HmiScreenItemData_11" at 836,128 size 203x35; TextOn 'Back'; TextOff 'Voyage A'
   Button "HmiScreenItemData_12" at 836,233 size 203x28; TextOn 'Back'; TextOff 'Pre Dwell Time'
   Button "HmiScreenItemData_13" at 836,267 size 203x28; TextOn 'Back'; TextOff 'De-Oxygenation Minimum Time'
   Button "HmiScreenItemData_43" at 836,335 size 203x28; TextOn 'Back'; TextOff 'Dwell Time'
   Button "HmiScreenItemData_44" at 836,369 size 203x28; TextOn 'Back'; TextOff 'Re-Oxygenation Time'
   Button "HmiScreenItemData_45" at 836,403 size 203x28; TextOn 'Back'; TextOff 'Post Dwell Time'
   IOField "I/O field_17" at 1060,169 size 79x28; Authorization "User administration"; FormatPattern 999; Unit  Hrs
      ProcessValue <- "2110_BTCS_CNTRL_DB_TOT_SEQ_HRS"
   Button "HmiScreenItemData_42" at 836,169 size 203x28; TextOn 'Back'; TextOff 'Total Treatment Time'
   Button "HmiScreenItemData_47" at 482,461 size 418x27; TextOn 'Back'; TextOff 'Automatic Ballast Tank Selection'
   Button "HmiScreenItemData_9" at 525,88 size 220x30; TextOn 'Back'; TextOff 'Pre Dwell Time Completed'
   Button "HmiScreenItemData_17" at 525,148 size 220x30; TextOn 'Back'; TextOff 'De-Oxygenation Completed'
   Button "HmiScreenItemData_38" at 525,178 size 220x30; TextOn 'Back'; TextOff 'Dwell Time Completed'
   Button "HmiScreenItemData_39" at 525,238 size 220x30; TextOn 'Back'; TextOff 'Re-Oxygenation Completed'
   Button "HmiScreenItemData_41" at 525,269 size 220x30; TextOn 'Back'; TextOff 'Post Dwell Time Completed'
   Button "HmiScreenItemData_46" at 525,118 size 220x30; TextOn 'Back'; TextOff 'Inert Gas Transfer Active'
   Button "HmiScreenItemData_48" at 525,208 size 220x30; TextOn 'Back'; TextOff 'Ambient Air Transfer Active'
   Button "HmiScreenItemData_52" at 525,118 size 220x30; TextOn 'Back'; TextOff 'IG Transfer Completed'
   Button "HmiScreenItemData_53" at 525,208 size 220x30; TextOn 'Back'; TextOff 'Ambient Air Transfer Completed'
   Button "HmiScreenItemData_3" at 1129,1 size 150x40; TextOn 'I&A Compressor Ok'; TextOff 'Back'
      on Release: function_efd93a16()
   TextField "Text field_11" at 1179,94 size 36x18; Text 'ETA'
   IOField "I/O field_16" at 1156,233 size 83x28; Authorization "User administration"; FormatPattern 999; Unit  min
      ProcessValue <- "2102_TIME_CALCS_DB_PRE_DWELL_MINS_RMNG"
   IOField "I/O field_18" at 1156,267 size 83x28; Authorization "User administration"; FormatPattern 999; Unit  min
   IOField "I/O field_19" at 1156,335 size 83x28; FormatPattern 999; Unit  min
      ProcessValue <- "2102_TIME_CALCS_DB_DWELL_MINS_RMNG"
   IOField "I/O field_20" at 1156,369 size 83x28; FormatPattern 999; Unit  min
      ProcessValue <- "2102_TIME_CALCS_DB_RE_OX_MINS_RMNG"
   IOField "I/O field_21" at 1156,403 size 83x28; FormatPattern 999; Unit  min
      ProcessValue <- "2102_TIME_CALCS_DB_POST_DWELL_MINS_RMNG"
   IOField "I/O field_22" at 1156,169 size 83x28; Authorization "User administration"; FormatPattern 999; Unit  Hrs
      ProcessValue <- "2110_BTCS_CNTRL_DB_RMNG_SEQ_HRS"
   Rectangle "Rectangle_25" at 281,165 size 179x59
      Visibility <- "2100_AUTO_SEQ_DB_SEQ_RNG"
   Button "HmiScreenItemData_4" at 282,172 size 150x47; TextOn 'Back'; TextOff 'Abort & Stop'; Authorization "Operating Mode"
      Appearance <- "2110_BTCS_CNTRL_DB_BTCS_STATE"
      on Release: function_efd93a16("BWTS Stop Confirm", 400, 200, -1, -1, 1)
      ObjectEnable <- "82_To_HMI_CRNT_MODE_GCU"
   Circle "Circle_9" at 453,125 size 29x29
      Appearance <- "2110_BTCS_CNTRL_DB_BTCS_STATE"
   Circle "Circle_1" at 453,181 size 29x29
      Appearance <- "2110_BTCS_CNTRL_DB_BTCS_STATE"
   TextField "Text field_60" at 936,698 size 290x35; Text 'SALINITY ACCEPTED'
      Visibility <- "2068_Sys_Status_Data_SAL_VALID"
   Circle "Circle_19" at 220,233 size 29x29
      Appearance <- "150_GCU_LCL_CNTRL_DB_LCL_CNTRL_ACTV"
   Circle "Circle_20" at 220,180 size 29x29
      Appearance <- "82_To_HMI_CRNT_MODE_GCU"
   Button "HmiScreenItemData_36" at 49,170 size 150x51; TextOn 'Back'; TextOff 'Manual'; Authorization "Operating Mode"
      on Press: function_b14e0dd5("80_From_HMI_Request_Manual", 0); ResetBit("150_GCU_LCL_CNTRL_DB_LCL_CNTRL_ACTV")
   Circle "Circle_21" at 220,126 size 29x29
      Appearance <- "82_To_HMI_CRNT_MODE_GCU"
   Button "HmiScreenItemData_37" at 49,116 size 150x51; TextOn 'Back'; TextOff 'Full Auto'; Authorization "Operating Mode"
      on Press: function_b14e0dd5("80_From_HMI_Request_Auto", 0); ResetBit("150_GCU_LCL_CNTRL_DB_LCL_CNTRL_ACTV")
   Button "HmiScreenItemData_49" at 49,225 size 150x51; TextOn 'Back'; TextOff 'Local Auto'; Authorization "User administration"
      on Press: InvertBit("150_GCU_LCL_CNTRL_DB_LCL_CNTRL_ACTV"); function_b14e0dd5("80_From_HMI_Request_Auto", 0); ResetBit("80_From_HMI_Request_Manual")
   Circle "Circle_22" at 220,126 size 29x29
      Visibility <- "150_GCU_LCL_CNTRL_DB_LCL_CNTRL_ACTV"
   Circle "Circle_30" at 220,233 size 29x29
      Visibility <- "82_To_HMI_CRNT_MODE_GCU"
   Button "Button_4" at 493,507 size 100x23; TextOff 'FPT'; Authorization "Operate"
      Appearance <- "504_Tank Grouping_DB2020_TANK ACTIV 1"
      on Press: function_b14e0dd5("504_Tank Grouping_DB2020_TANK ACTIV 1", 0)
   IOField "I/O field_1" at 1040,301 size 79x28; Authorization "Commissioning"; FormatPattern 999; Unit  Hrs
      ProcessValue <- "2110_BTCS_CNTRL_DB_DE_OX_SP_HRS"
   Button "HmiScreenItemData_6" at 836,301 size 203x28; TextOn 'Back'; TextOff 'De-Oxygenation Setpoint Time'
   Rectangle "Rectangle_21" at 917,659 size 327x40
      Appearance <- "2068_Sys_Status_Data_SAL_VALID"
   TextField "Text field_48" at 916,664 size 128x30; Text 'Salinity Value:'
   IOField "I/O field_31" at 1036,664 size 74x30; FormatPattern 99.9; Unit psu
      ProcessValue <- "80_From_HMI_SAL_VALUE"
   Button "HmiScreenItemData_35" at 1108,664 size 135x30; TextOn 'Back'; TextOff 'Confirm Salinity'
      on Release: function_efd93a16("Salinity - Acceptance", 0, 0, 1, 3, 1)
   Group "Group_18" at 921,659 size 322x40
   Group "Group" at 916,659 size 327x40; Authorization "Operate"
   Button "HmiScreenItemData_7" at 1156,85 size 83x35; TextOn 'CONTINUE'; TextOff 'Continue'; Authorization "Operating Mode"
      on Press: InvertBit("80_From_HMI_TIMER RST Supres")
      Appearance <- "80_From_HMI_TIMER RST Supres"
   IOField "I/O field_25" at 1040,201 size 79x28; Authorization "User administration"; FormatPattern 999.9; Unit  Hrs
      ProcessValue <- "504_Tank Grouping_DB2020_Sequence Time m Offset_Int"
   Button "HmiScreenItemData_2" at 836,201 size 203x28; TextOn 'Back'; TextOff 'Differential Treatment Time'
   IOField "I/O field_3" at 1156,201 size 83x28; Authorization "User administration"; FormatPattern 999; Unit  min
      ProcessValue <- "504_Tank Grouping_DB2020_Diff Time Remain"
   Button "Button_1" at 817,594 size 79x32; TextOff '3'; Authorization "Operate"
      Appearance <- "504_Tank Grouping_DB2020_GROUP ACTIVE INT 3"
      on Press: function_b14e0dd5("504_Tank Grouping_DB2020_GROUP ACTIV 3", 0)
   Button "Button_2" at 817,628 size 79x32; TextOff '4'; Authorization "Operate"
      Appearance <- "504_Tank Grouping_DB2020_GROUP ACTIVE INT 4"
      on Press: function_b14e0dd5("504_Tank Grouping_DB2020_GROUP ACTIV 4", 0)
   Button "Button_10" at 818,662 size 79x32; TextOff '5'; Authorization "Operate"
      Appearance <- "504_Tank Grouping_DB2020_GROUP ACTIVE INT 5"
      on Press: function_b14e0dd5("504_Tank Grouping_DB2020_GROUP ACTIV 5", 0)
   Button "Button_11" at 818,696 size 79x32; TextOff '6'; Authorization "Operate"
      Appearance <- "504_Tank Grouping_DB2020_GROUP ACTIVE INT 6"
      on Press: function_b14e0dd5("504_Tank Grouping_DB2020_GROUP ACTIV 6", 0)
   Button "Button_12" at 818,731 size 79x32; TextOff '7'; Authorization "Operate"
      Appearance <- "504_Tank Grouping_DB2020_GROUP ACTIVE INT 7"
      on Press: function_b14e0dd5("504_Tank Grouping_DB2020_GROUP ACTIV 7", 0)